// TIA Portal project "CLU" (V13) (continued)
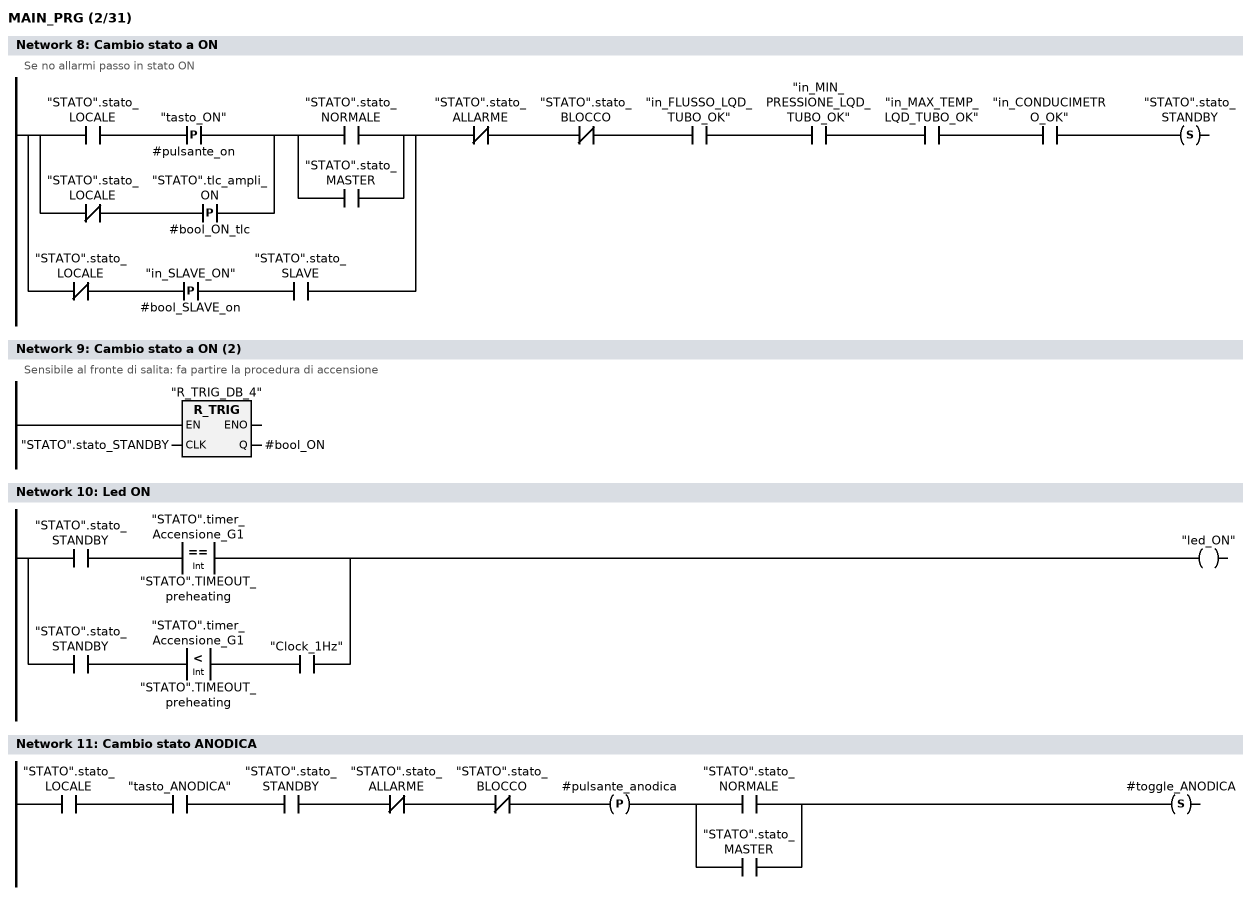
   RUNG wire#powerrail
      Contact( "STATO".stato_LOCALE )
      P_Contact(operand := "tasto_ON", bit := #pulsante_on)
      wire#w1
      Contact( "STATO".stato_NORMALE )
      wire#w2
      I_Contact( "STATO".stato_ALLARME )
      I_Contact( "STATO".stato_BLOCCO )
      Contact( "in_FLUSSO_LQD_TUBO_OK" )
      Contact( "in_MIN_PRESSIONE_LQD_TUBO_OK" )
      Contact( "in_MAX_TEMP_LQD_TUBO_OK" )
      Contact( "in_CONDUCIMETRO_OK" )
      S_Coil( "STATO".stato_STANDBY )
   END_RUNG
   RUNG wire#powerrail
      I_Contact( "STATO".stato_LOCALE )
      P_Contact(operand := "STATO".tlc_ampli_ON, bit := #bool_ON_tlc)
   END_RUNG wire#w1
   RUNG wire#w1
      Contact( "STATO".stato_MASTER )
   END_RUNG wire#w2
   RUNG wire#powerrail
      I_Contact( "STATO".stato_LOCALE )
      P_Contact(operand := "in_SLAVE_ON", bit := #bool_SLAVE_on)
      Contact( "STATO".stato_SLAVE )
   END_RUNG wire#w2
   // the same network as SCL:
   #_w1 := "STATO".stato_LOCALE AND "tasto_ON" AND NOT #pulsante_on;   // rising edge of "tasto_ON"
   #pulsante_on := "tasto_ON";
   #_w2 := NOT "STATO".stato_LOCALE AND "STATO".tlc_ampli_ON AND NOT #bool_ON_tlc;   // rising edge of "STATO".tlc_ampli_ON
   #bool_ON_tlc := "STATO".tlc_ampli_ON;
   #_w3 := NOT "STATO".stato_LOCALE AND "in_SLAVE_ON" AND NOT #bool_SLAVE_on;   // rising edge of "in_SLAVE_ON"
   #bool_SLAVE_on := "in_SLAVE_ON";
   IF (((#_w1 OR #_w2) AND ("STATO".stato_NORMALE OR "STATO".stato_MASTER)) OR (#_w3 AND "STATO".stato_SLAVE)) AND NOT "STATO".stato_ALLARME AND NOT "STATO".stato_BLOCCO AND "in_FLUSSO_LQD_TUBO_OK" AND "in_MIN_PRESSIONE_LQD_TUBO_OK" AND "in_MAX_TEMP_LQD_TUBO_OK" AND "in_CONDUCIMETRO_OK" THEN
       "STATO".stato_STANDBY := TRUE;
   END_IF;
END_REGION

REGION Network 9: Cambio stato a ON (2)
   // Sensibile al fronte di salita: fa partire la procedura di accensione
   "R_TRIG_DB_4"(CLK := "STATO".stato_STANDBY, Q => #bool_ON);   // R_TRIG
END_REGION

REGION Network 10: Led ON
   RUNG wire#powerrail
      Contact( "STATO".stato_STANDBY )
      { S7_Templates := "SrcType := Int" } EQ_Contact(in1 := "STATO".timer_Accensione_G1, in2 := "STATO".TIMEOUT_preheating)
      wire#w1
      Coil( "led_ON" )
   END_RUNG
   RUNG wire#powerrail
      Contact( "STATO".stato_STANDBY )
      { S7_Templates := "SrcType := Int" } LT_Contact(in1 := "STATO".timer_Accensione_G1, in2 := "STATO".TIMEOUT_preheating)
      Contact( "Clock_1Hz" )
   END_RUNG wire#w1
   // the same network as SCL:
   "led_ON" := ("STATO".stato_STANDBY AND ("STATO".timer_Accensione_G1 = "STATO".TIMEOUT_preheating)) OR ("STATO".stato_STANDBY AND ("STATO".timer_Accensione_G1 < "STATO".TIMEOUT_preheating) AND "Clock_1Hz");
END_REGION

REGION Network 11: Cambio stato ANODICA
   RUNG wire#powerrail
      Contact( "STATO".stato_LOCALE )
      Contact( "tasto_ANODICA" )
      Contact( "STATO".stato_STANDBY )
      I_Contact( "STATO".stato_ALLARME )
      I_Contact( "STATO".stato_BLOCCO )
      P_Trig( #pulsante_anodica )
      wire#w1
      Contact( "STATO".stato_NORMALE )
      wire#w2
      S_Coil( #toggle_ANODICA )
   END_RUNG
   RUNG wire#w1
      Contact( "STATO".stato_MASTER )
   END_RUNG wire#w2
   // the same network as SCL:
   #_w1 := "STATO".stato_LOCALE AND "tasto_ANODICA" AND "STATO".stato_STANDBY AND NOT "STATO".stato_ALLARME AND NOT "STATO".stato_BLOCCO;
   #_w2 := #_w1 AND NOT #pulsante_anodica;   // rising edge
   #pulsante_anodica := #_w1;
   IF #_w2 AND ("STATO".stato_NORMALE OR "STATO".stato_MASTER) THEN #toggle_ANODICA := TRUE; END_IF;
END_REGION

REGION Network 12: ANODICA ON
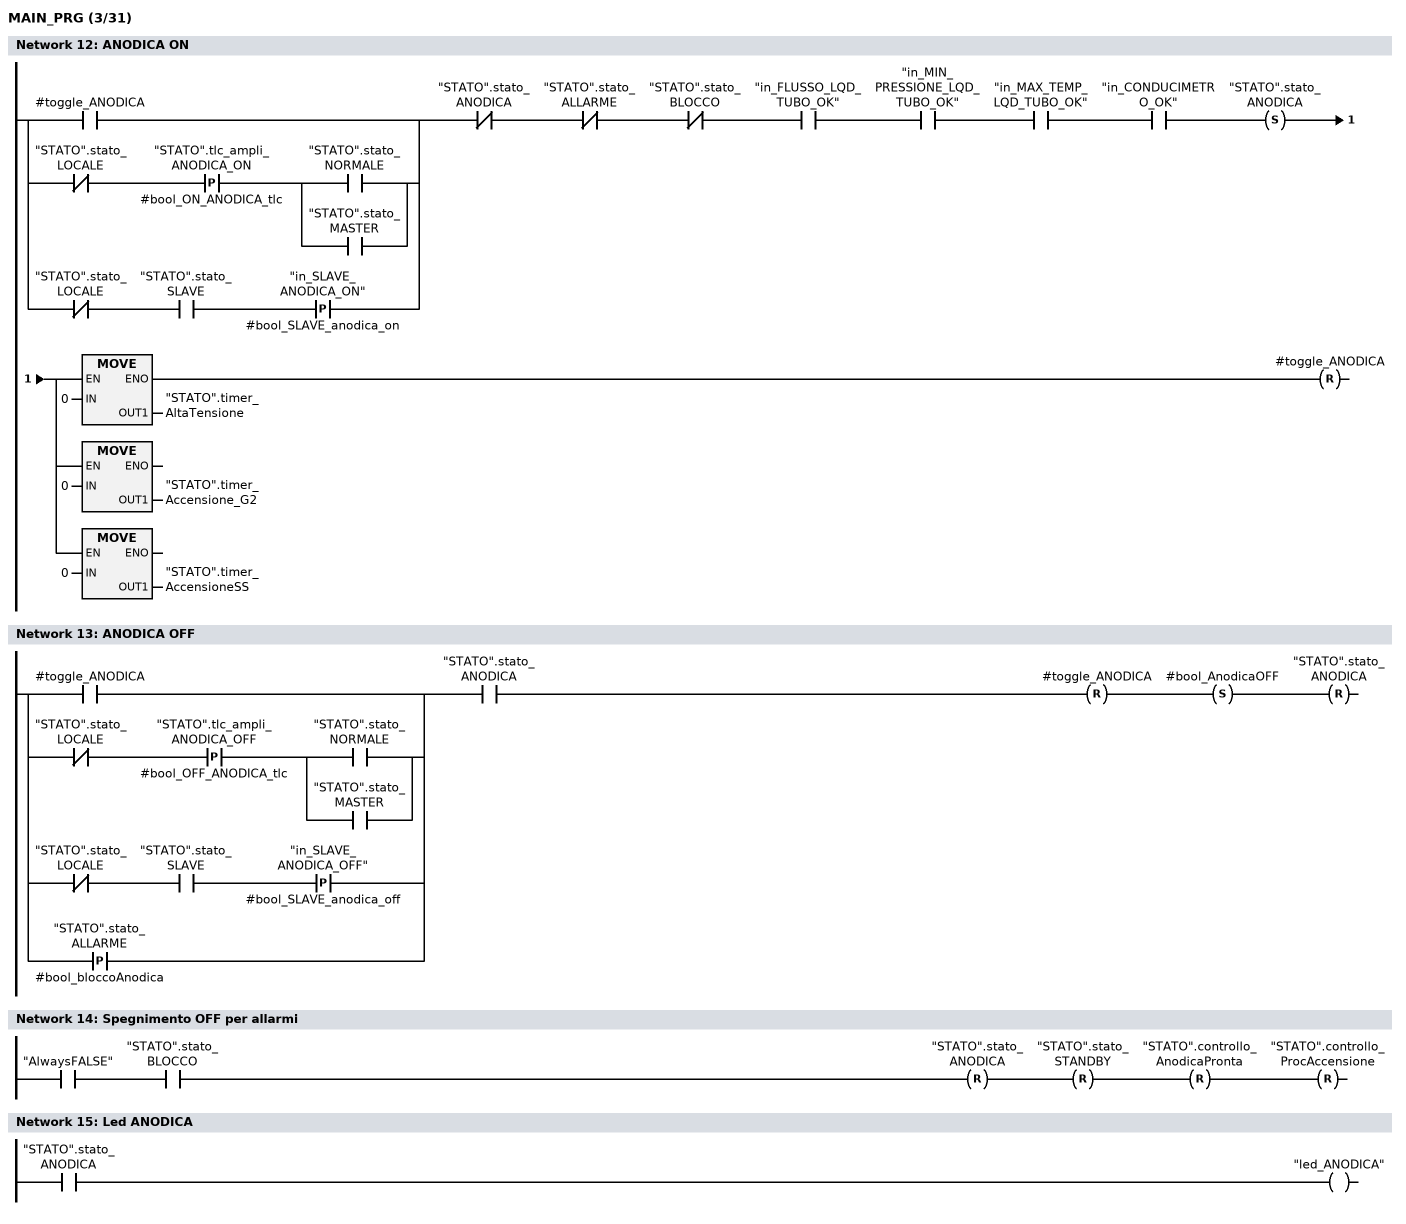
   RUNG wire#powerrail
      Contact( #toggle_ANODICA )
      wire#w1
      I_Contact( "STATO".stato_ANODICA )
      I_Contact( "STATO".stato_ALLARME )
      I_Contact( "STATO".stato_BLOCCO )
      Contact( "in_FLUSSO_LQD_TUBO_OK" )
      Contact( "in_MIN_PRESSIONE_LQD_TUBO_OK" )
      Contact( "in_MAX_TEMP_LQD_TUBO_OK" )
      Contact( "in_CONDUCIMETRO_OK" )
      S_Coil( "STATO".stato_ANODICA )
      wire#w3
      Move(in := 0, out1 => "STATO".timer_AltaTensione)
      R_Coil( #toggle_ANODICA )
   END_RUNG
   RUNG wire#powerrail
      I_Contact( "STATO".stato_LOCALE )
      P_Contact(operand := "STATO".tlc_ampli_ANODICA_ON, bit := #bool_ON_ANODICA_tlc)
      wire#w2
      Contact( "STATO".stato_NORMALE )
   END_RUNG wire#w1
   RUNG wire#w2
      Contact( "STATO".stato_MASTER )
   END_RUNG wire#w1
   RUNG wire#powerrail
      I_Contact( "STATO".stato_LOCALE )
      Contact( "STATO".stato_SLAVE )
      P_Contact(operand := "in_SLAVE_ANODICA_ON", bit := #bool_SLAVE_anodica_on)
   END_RUNG wire#w1
   RUNG wire#w3
      Move(in := 0, out1 => "STATO".timer_Accensione_G2)
   END_RUNG
   RUNG wire#w3
      Move(in := 0, out1 => "STATO".timer_AccensioneSS)
   END_RUNG
   // the same network as SCL:
   #_w1 := NOT "STATO".stato_LOCALE AND "STATO".tlc_ampli_ANODICA_ON AND NOT #bool_ON_ANODICA_tlc;   // rising edge of "STATO".tlc_ampli_ANODICA_ON
   #bool_ON_ANODICA_tlc := "STATO".tlc_ampli_ANODICA_ON;
   #_w2 := NOT "STATO".stato_LOCALE AND "STATO".stato_SLAVE AND "in_SLAVE_ANODICA_ON" AND NOT #bool_SLAVE_anodica_on;   // rising edge of "in_SLAVE_ANODICA_ON"
   #bool_SLAVE_anodica_on := "in_SLAVE_ANODICA_ON";
   #_w3 := (#toggle_ANODICA OR (#_w1 AND ("STATO".stato_NORMALE OR "STATO".stato_MASTER)) OR #_w2) AND NOT "STATO".stato_ANODICA AND NOT "STATO".stato_ALLARME AND NOT "STATO".stato_BLOCCO AND "in_FLUSSO_LQD_TUBO_OK" AND "in_MIN_PRESSIONE_LQD_TUBO_OK" AND "in_MAX_TEMP_LQD_TUBO_OK" AND "in_CONDUCIMETRO_OK";
   IF #_w3 THEN
       "STATO".stato_ANODICA := TRUE;
       "STATO".timer_AltaTensione := 0;
       #toggle_ANODICA := FALSE;
       "STATO".timer_Accensione_G2 := 0;
       "STATO".timer_AccensioneSS := 0;
   END_IF;
END_REGION

REGION Network 13: ANODICA OFF
   RUNG wire#powerrail
      Contact( #toggle_ANODICA )
      wire#w1
      Contact( "STATO".stato_ANODICA )
      R_Coil( #toggle_ANODICA )
      S_Coil( #bool_AnodicaOFF )
      R_Coil( "STATO".stato_ANODICA )
   END_RUNG
   RUNG wire#powerrail
      I_Contact( "STATO".stato_LOCALE )
      P_Contact(operand := "STATO".tlc_ampli_ANODICA_OFF, bit := #bool_OFF_ANODICA_tlc)
      wire#w2
      Contact( "STATO".stato_NORMALE )
   END_RUNG wire#w1
   RUNG wire#w2
      Contact( "STATO".stato_MASTER )
   END_RUNG wire#w1
   RUNG wire#powerrail
      I_Contact( "STATO".stato_LOCALE )
      Contact( "STATO".stato_SLAVE )
      P_Contact(operand := "in_SLAVE_ANODICA_OFF", bit := #bool_SLAVE_anodica_off)
   END_RUNG wire#w1
   RUNG wire#powerrail
      P_Contact(operand := "STATO".stato_ALLARME, bit := #bool_bloccoAnodica)
   END_RUNG wire#w1
   // the same network as SCL:
   #_w1 := NOT "STATO".stato_LOCALE AND "STATO".tlc_ampli_ANODICA_OFF AND NOT #bool_OFF_ANODICA_tlc;   // rising edge of "STATO".tlc_ampli_ANODICA_OFF
   #bool_OFF_ANODICA_tlc := "STATO".tlc_ampli_ANODICA_OFF;
   #_w2 := NOT "STATO".stato_LOCALE AND "STATO".stato_SLAVE AND "in_SLAVE_ANODICA_OFF" AND NOT #bool_SLAVE_anodica_off;   // rising edge of "in_SLAVE_ANODICA_OFF"
   #bool_SLAVE_anodica_off := "in_SLAVE_ANODICA_OFF";
   #_w3 := "STATO".stato_ALLARME AND NOT #bool_bloccoAnodica;   // rising edge of "STATO".stato_ALLARME
   #bool_bloccoAnodica := "STATO".stato_ALLARME;
   #_w4 := (#toggle_ANODICA OR (#_w1 AND ("STATO".stato_NORMALE OR "STATO".stato_MASTER)) OR #_w2 OR #_w3) AND "STATO".stato_ANODICA;
   IF #_w4 THEN
       #toggle_ANODICA := FALSE;
       #bool_AnodicaOFF := TRUE;
       "STATO".stato_ANODICA := FALSE;
   END_IF;
END_REGION

REGION Network 14: Spegnimento OFF per allarmi
   RUNG wire#powerrail
      Contact( "AlwaysFALSE" )
      Contact( "STATO".stato_BLOCCO )
      R_Coil( "STATO".stato_ANODICA )
      R_Coil( "STATO".stato_STANDBY )
      R_Coil( "STATO".controllo_AnodicaPronta )
      R_Coil( "STATO".controllo_ProcAccensione )
   END_RUNG
   // the same network as SCL:
   IF "AlwaysFALSE" AND "STATO".stato_BLOCCO THEN
       "STATO".stato_ANODICA := FALSE;
       "STATO".stato_STANDBY := FALSE;
       "STATO".controllo_AnodicaPronta := FALSE;
       "STATO".controllo_ProcAccensione := FALSE;
   END_IF;
END_REGION

REGION Network 15: Led ANODICA
   RUNG wire#powerrail
      Contact( "STATO".stato_ANODICA )
      Coil( "led_ANODICA" )
   END_RUNG
   // the same network as SCL:
   "led_ANODICA" := "STATO".stato_ANODICA;
END_REGION

REGION Network 16: Cambio a modo CW /Pulsed
   // Non applicabile se l'Anodica è attiva
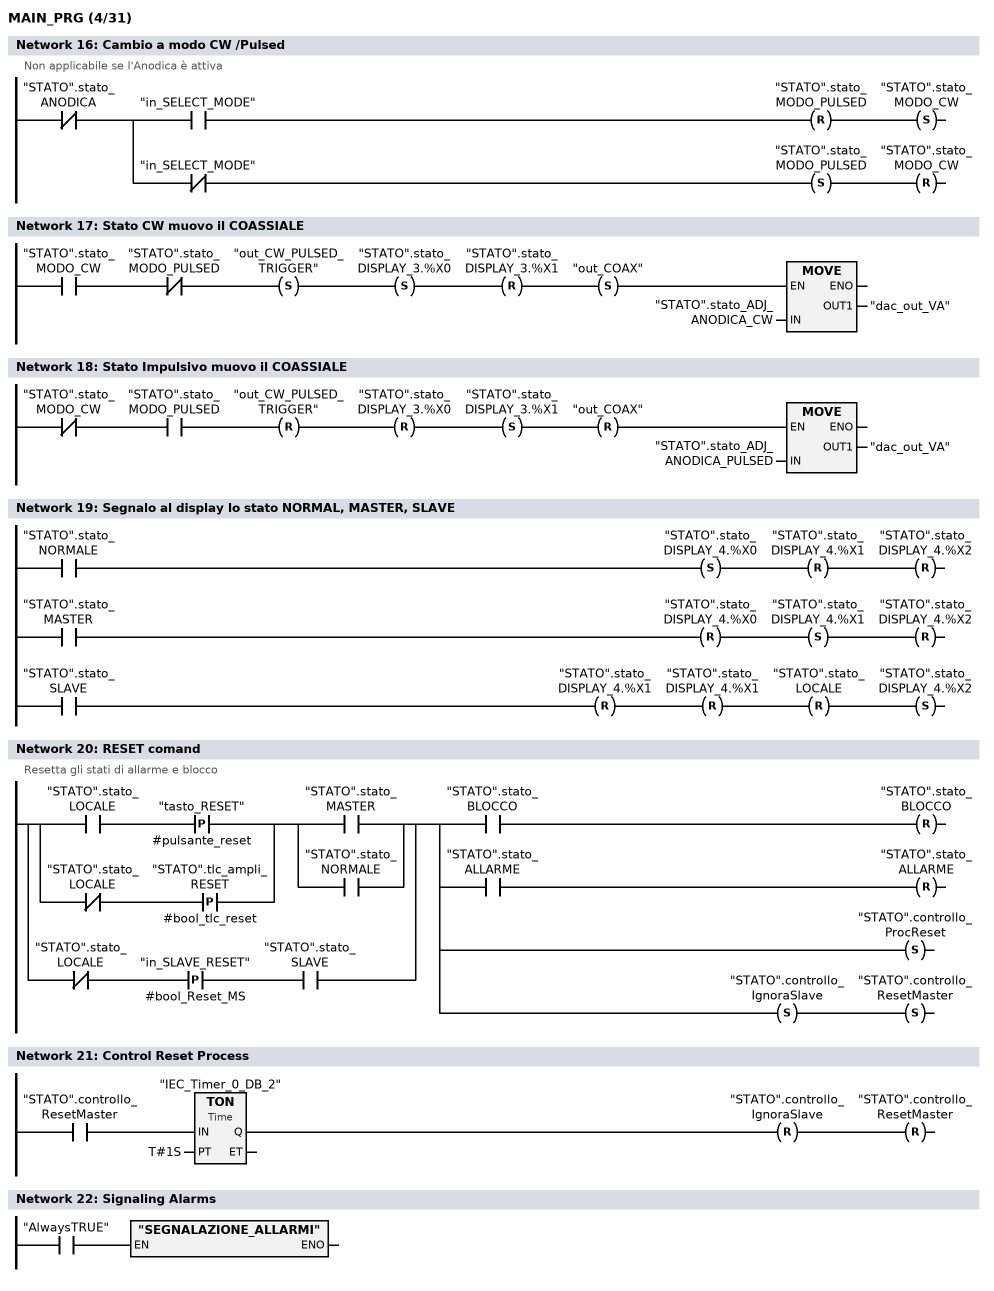
   RUNG wire#powerrail
      I_Contact( "STATO".stato_ANODICA )
      wire#w1
      Contact( "in_SELECT_MODE" )
      R_Coil( "STATO".stato_MODO_PULSED )
      S_Coil( "STATO".stato_MODO_CW )
   END_RUNG
   RUNG wire#w1
      I_Contact( "in_SELECT_MODE" )
      S_Coil( "STATO".stato_MODO_PULSED )
      R_Coil( "STATO".stato_MODO_CW )
   END_RUNG
   // the same network as SCL:
   #_w1 := NOT "STATO".stato_ANODICA;
   IF #_w1 AND "in_SELECT_MODE" THEN
       "STATO".stato_MODO_PULSED := FALSE;
       "STATO".stato_MODO_CW := TRUE;
   END_IF;
   IF #_w1 AND NOT "in_SELECT_MODE" THEN
       "STATO".stato_MODO_PULSED := TRUE;
       "STATO".stato_MODO_CW := FALSE;
   END_IF;
END_REGION

REGION Network 17: Stato CW muovo il COASSIALE
   RUNG wire#powerrail
      Contact( "STATO".stato_MODO_CW )
      I_Contact( "STATO".stato_MODO_PULSED )
      S_Coil( "out_CW_PULSED_TRIGGER" )
      S_Coil( "STATO".stato_DISPLAY_3.%X0 )
      R_Coil( "STATO".stato_DISPLAY_3.%X1 )
      S_Coil( "out_COAX" )
      Move(in := "STATO".stato_ADJ_ANODICA_CW, out1 => "dac_out_VA")
   END_RUNG
   // the same network as SCL:
   IF "STATO".stato_MODO_CW AND NOT "STATO".stato_MODO_PULSED THEN
       "out_CW_PULSED_TRIGGER" := TRUE;
       "STATO".stato_DISPLAY_3.%X0 := TRUE;
       "STATO".stato_DISPLAY_3.%X1 := FALSE;
       "out_COAX" := TRUE;
       "dac_out_VA" := "STATO".stato_ADJ_ANODICA_CW;
   END_IF;
END_REGION

REGION Network 18: Stato Impulsivo muovo il COASSIALE
   RUNG wire#powerrail
      I_Contact( "STATO".stato_MODO_CW )
      Contact( "STATO".stato_MODO_PULSED )
      R_Coil( "out_CW_PULSED_TRIGGER" )
      R_Coil( "STATO".stato_DISPLAY_3.%X0 )
      S_Coil( "STATO".stato_DISPLAY_3.%X1 )
      R_Coil( "out_COAX" )
      Move(in := "STATO".stato_ADJ_ANODICA_PULSED, out1 => "dac_out_VA")
   END_RUNG
   // the same network as SCL:
   IF NOT "STATO".stato_MODO_CW AND "STATO".stato_MODO_PULSED THEN
       "out_CW_PULSED_TRIGGER" := FALSE;
       "STATO".stato_DISPLAY_3.%X0 := FALSE;
       "STATO".stato_DISPLAY_3.%X1 := TRUE;
       "out_COAX" := FALSE;
       "dac_out_VA" := "STATO".stato_ADJ_ANODICA_PULSED;
   END_IF;
END_REGION

REGION Network 19: Segnalo al display lo stato NORMAL, MASTER, SLAVE
   RUNG wire#powerrail
      Contact( "STATO".stato_NORMALE )
      S_Coil( "STATO".stato_DISPLAY_4.%X0 )
      R_Coil( "STATO".stato_DISPLAY_4.%X1 )
      R_Coil( "STATO".stato_DISPLAY_4.%X2 )
   END_RUNG
   RUNG wire#powerrail
      Contact( "STATO".stato_MASTER )
      R_Coil( "STATO".stato_DISPLAY_4.%X0 )
      S_Coil( "STATO".stato_DISPLAY_4.%X1 )
      R_Coil( "STATO".stato_DISPLAY_4.%X2 )
   END_RUNG
   RUNG wire#powerrail
      Contact( "STATO".stato_SLAVE )
      R_Coil( "STATO".stato_DISPLAY_4.%X1 )
      R_Coil( "STATO".stato_DISPLAY_4.%X1 )
      R_Coil( "STATO".stato_LOCALE )
      S_Coil( "STATO".stato_DISPLAY_4.%X2 )
   END_RUNG
   // the same network as SCL:
   IF "STATO".stato_NORMALE THEN
       "STATO".stato_DISPLAY_4.%X0 := TRUE;
       "STATO".stato_DISPLAY_4.%X1 := FALSE;
       "STATO".stato_DISPLAY_4.%X2 := FALSE;
   END_IF;
   IF "STATO".stato_MASTER THEN
       "STATO".stato_DISPLAY_4.%X0 := FALSE;
       "STATO".stato_DISPLAY_4.%X1 := TRUE;
       "STATO".stato_DISPLAY_4.%X2 := FALSE;
   END_IF;
   IF "STATO".stato_SLAVE THEN
       "STATO".stato_DISPLAY_4.%X1 := FALSE;
       "STATO".stato_DISPLAY_4.%X1 := FALSE;
       "STATO".stato_LOCALE := FALSE;
       "STATO".stato_DISPLAY_4.%X2 := TRUE;
   END_IF;
END_REGION

REGION Network 20: RESET comand
   // Resetta gli stati di allarme e blocco
   RUNG wire#powerrail
      Contact( "STATO".stato_LOCALE )
      P_Contact(operand := "tasto_RESET", bit := #pulsante_reset)
      wire#w1
      Contact( "STATO".stato_MASTER )
      wire#w2
      Contact( "STATO".stato_BLOCCO )
      R_Coil( "STATO".stato_BLOCCO )
   END_RUNG
   RUNG wire#powerrail
      I_Contact( "STATO".stato_LOCALE )
      P_Contact(operand := "STATO".tlc_ampli_RESET, bit := #bool_tlc_reset)
   END_RUNG wire#w1
   RUNG wire#w1
      Contact( "STATO".stato_NORMALE )
   END_RUNG wire#w2
   RUNG wire#powerrail
      I_Contact( "STATO".stato_LOCALE )
      P_Contact(operand := "in_SLAVE_RESET", bit := #bool_Reset_MS)
      Contact( "STATO".stato_SLAVE )
   END_RUNG wire#w2
   RUNG wire#w2
      Contact( "STATO".stato_ALLARME )
      R_Coil( "STATO".stato_ALLARME )
   END_RUNG
   RUNG wire#w2
      S_Coil( "STATO".controllo_ProcReset )
   END_RUNG
   RUNG wire#w2
      S_Coil( "STATO".controllo_IgnoraSlave )
      S_Coil( "STATO".controllo_ResetMaster )
   END_RUNG
   // the same network as SCL:
   #_w1 := "STATO".stato_LOCALE AND "tasto_RESET" AND NOT #pulsante_reset;   // rising edge of "tasto_RESET"
   #pulsante_reset := "tasto_RESET";
   #_w2 := NOT "STATO".stato_LOCALE AND "STATO".tlc_ampli_RESET AND NOT #bool_tlc_reset;   // rising edge of "STATO".tlc_ampli_RESET
   #bool_tlc_reset := "STATO".tlc_ampli_RESET;
   #_w3 := NOT "STATO".stato_LOCALE AND "in_SLAVE_RESET" AND NOT #bool_Reset_MS;   // rising edge of "in_SLAVE_RESET"
   #bool_Reset_MS := "in_SLAVE_RESET";
   #_w4 := ((#_w1 OR #_w2) AND ("STATO".stato_MASTER OR "STATO".stato_NORMALE)) OR (#_w3 AND "STATO".stato_SLAVE);
   IF #_w4 AND "STATO".stato_BLOCCO THEN "STATO".stato_BLOCCO := FALSE; END_IF;
   IF #_w4 AND "STATO".stato_ALLARME THEN "STATO".stato_ALLARME := FALSE; END_IF;
   IF #_w4 THEN
       "STATO".controllo_ProcReset := TRUE;
       "STATO".controllo_IgnoraSlave := TRUE;
       "STATO".controllo_ResetMaster := TRUE;
   END_IF;
END_REGION

REGION Network 21: Control Reset Process
   "IEC_Timer_0_DB_2".TON(IN := "STATO".controllo_ResetMaster, PT := T#1S);
   IF "IEC_Timer_0_DB_2".Q THEN
       "STATO".controllo_IgnoraSlave := FALSE;
       "STATO".controllo_ResetMaster := FALSE;
   END_IF;
END_REGION

REGION Network 22: Signaling Alarms
   RUNG wire#powerrail
      Contact( "AlwaysTRUE" )
      "SEGNALAZIONE_ALLARMI"()
   END_RUNG
   // the same network as SCL:
   IF "AlwaysTRUE" THEN "SEGNALAZIONE_ALLARMI"(); END_IF;
END_REGION

REGION Network 23: Erasing Alarms
   // In seguito ad un reset.
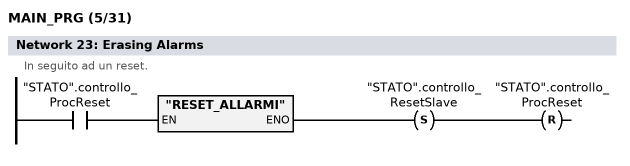
   RUNG wire#powerrail
      Contact( "STATO".controllo_ProcReset )
      "RESET_ALLARMI"()
      S_Coil( "STATO".controllo_ResetSlave )
      R_Coil( "STATO".controllo_ProcReset )
   END_RUNG
   // the same network as SCL:
   "RESET_ALLARMI"(EN := "STATO".controllo_ProcReset, ENO => #_w1);
   IF #_w1 THEN
       "STATO".controllo_ResetSlave := TRUE;
       "STATO".controllo_ProcReset := FALSE;
   END_IF;
END_REGION

REGION Network 24: ALARM STATE
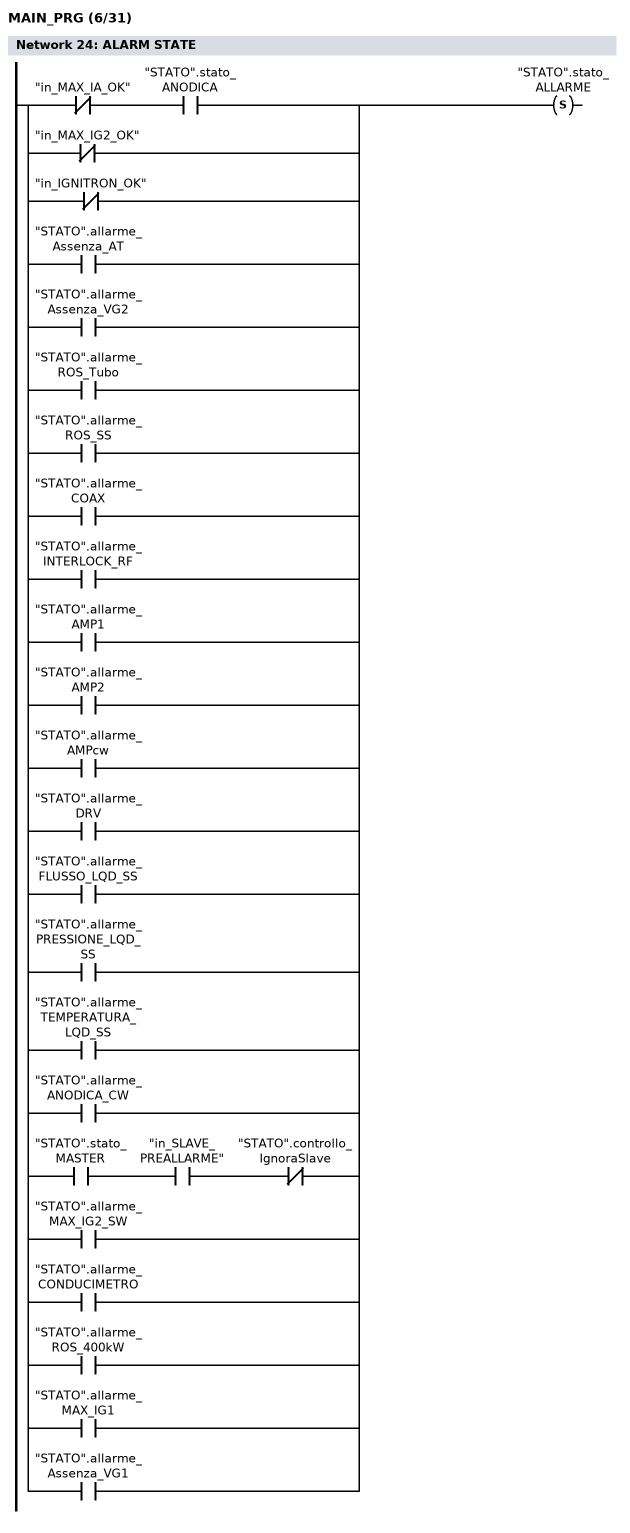
   RUNG wire#powerrail
      I_Contact( "in_MAX_IA_OK" )
      Contact( "STATO".stato_ANODICA )
      wire#w1
      S_Coil( "STATO".stato_ALLARME )
   END_RUNG
   RUNG wire#powerrail
      I_Contact( "in_MAX_IG2_OK" )
   END_RUNG wire#w1
   RUNG wire#powerrail
      I_Contact( "in_IGNITRON_OK" )
   END_RUNG wire#w1
   RUNG wire#powerrail
      Contact( "STATO".allarme_Assenza_AT )
   END_RUNG wire#w1
   RUNG wire#powerrail
      Contact( "STATO".allarme_Assenza_VG2 )
   END_RUNG wire#w1
   RUNG wire#powerrail
      Contact( "STATO".allarme_ROS_Tubo )
   END_RUNG wire#w1
   RUNG wire#powerrail
      Contact( "STATO".allarme_ROS_SS )
   END_RUNG wire#w1
   RUNG wire#powerrail
      Contact( "STATO".allarme_COAX )
   END_RUNG wire#w1
   RUNG wire#powerrail
      Contact( "STATO".allarme_INTERLOCK_RF )
   END_RUNG wire#w1
   RUNG wire#powerrail
      Contact( "STATO".allarme_AMP1 )
   END_RUNG wire#w1
   RUNG wire#powerrail
      Contact( "STATO".allarme_AMP2 )
   END_RUNG wire#w1
   RUNG wire#powerrail
      Contact( "STATO".allarme_AMPcw )
   END_RUNG wire#w1
   RUNG wire#powerrail
      Contact( "STATO".allarme_DRV )
   END_RUNG wire#w1
   RUNG wire#powerrail
      Contact( "STATO".allarme_FLUSSO_LQD_SS )
   END_RUNG wire#w1
   RUNG wire#powerrail
      Contact( "STATO".allarme_PRESSIONE_LQD_SS )
   END_RUNG wire#w1
   RUNG wire#powerrail
      Contact( "STATO".allarme_TEMPERATURA_LQD_SS )
   END_RUNG wire#w1
   RUNG wire#powerrail
      Contact( "STATO".allarme_ANODICA_CW )
   END_RUNG wire#w1
   RUNG wire#powerrail
      Contact( "STATO".stato_MASTER )
      Contact( "in_SLAVE_PREALLARME" )
      I_Contact( "STATO".controllo_IgnoraSlave )
   END_RUNG wire#w1
   RUNG wire#powerrail
      Contact( "STATO".allarme_MAX_IG2_SW )
   END_RUNG wire#w1
   RUNG wire#powerrail
      Contact( "STATO".allarme_CONDUCIMETRO )
   END_RUNG wire#w1
   RUNG wire#powerrail
      Contact( "STATO".allarme_ROS_400kW )
   END_RUNG wire#w1
   RUNG wire#powerrail
      Contact( "STATO".allarme_MAX_IG1 )
   END_RUNG wire#w1
   RUNG wire#powerrail
      Contact( "STATO".allarme_Assenza_VG1 )
   END_RUNG wire#w1
   // the same network as SCL:
   IF (NOT "in_MAX_IA_OK" AND "STATO".stato_ANODICA) OR NOT "in_MAX_IG2_OK" OR NOT "in_IGNITRON_OK" OR "STATO".allarme_Assenza_AT OR "STATO".allarme_Assenza_VG2 OR "STATO".allarme_ROS_Tubo OR "STATO".allarme_ROS_SS OR "STATO".allarme_COAX OR "STATO".allarme_INTERLOCK_RF OR "STATO".allarme_AMP1 OR "STATO".allarme_AMP2 OR "STATO".allarme_AMPcw OR "STATO".allarme_DRV OR "STATO".allarme_FLUSSO_LQD_SS OR "STATO".allarme_PRESSIONE_LQD_SS OR "STATO".allarme_TEMPERATURA_LQD_SS OR "STATO".allarme_ANODICA_CW OR ("STATO".stato_MASTER AND "in_SLAVE_PREALLARME" AND NOT "STATO".controllo_IgnoraSlave) OR "STATO".allarme_MAX_IG2_SW OR "STATO".allarme_CONDUCIMETRO OR "STATO".allarme_ROS_400kW OR "STATO".allarme_MAX_IG1 OR "STATO".allarme_Assenza_VG1 THEN
       "STATO".stato_ALLARME := TRUE;
   END_IF;
END_REGION

REGION Network 25: FAULT STATE
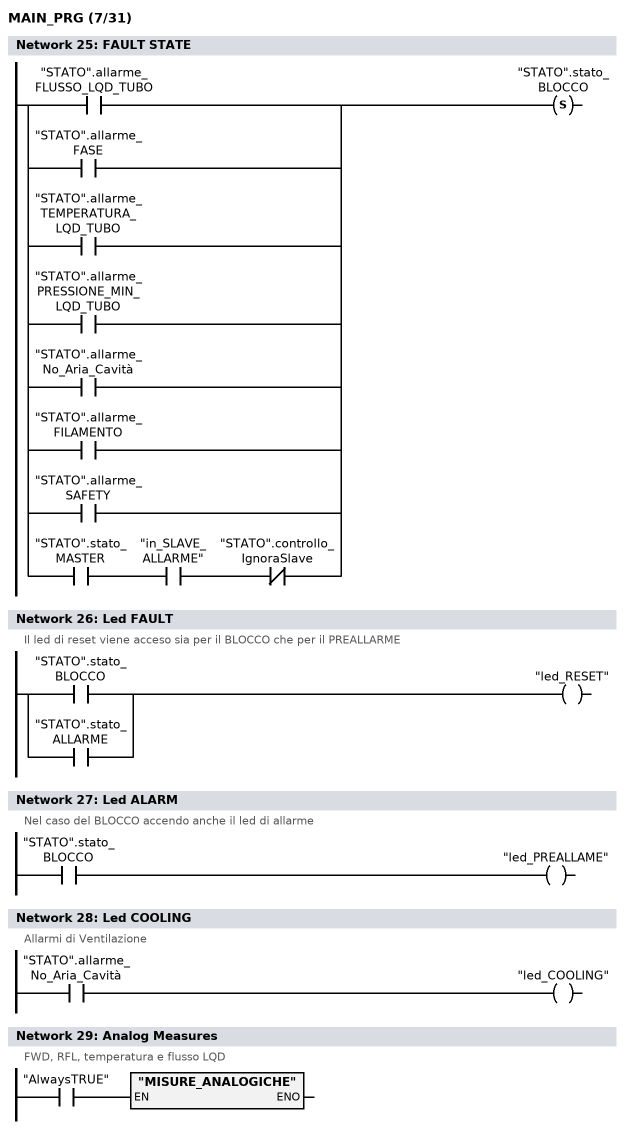
   RUNG wire#powerrail
      Contact( "STATO".allarme_FLUSSO_LQD_TUBO )
      wire#w1
      S_Coil( "STATO".stato_BLOCCO )
   END_RUNG
   RUNG wire#powerrail
      Contact( "STATO".allarme_FASE )
   END_RUNG wire#w1
   RUNG wire#powerrail
      Contact( "STATO".allarme_TEMPERATURA_LQD_TUBO )
   END_RUNG wire#w1
   RUNG wire#powerrail
      Contact( "STATO".allarme_PRESSIONE_MIN_LQD_TUBO )
   END_RUNG wire#w1
   RUNG wire#powerrail
      Contact( "STATO".allarme_No_Aria_Cavità )
   END_RUNG wire#w1
   RUNG wire#powerrail
      Contact( "STATO".allarme_FILAMENTO )
   END_RUNG wire#w1
   RUNG wire#powerrail
      Contact( "STATO".allarme_SAFETY )
   END_RUNG wire#w1
   RUNG wire#powerrail
      Contact( "STATO".stato_MASTER )
      Contact( "in_SLAVE_ALLARME" )
      I_Contact( "STATO".controllo_IgnoraSlave )
   END_RUNG wire#w1
   // the same network as SCL:
   IF "STATO".allarme_FLUSSO_LQD_TUBO OR "STATO".allarme_FASE OR "STATO".allarme_TEMPERATURA_LQD_TUBO OR "STATO".allarme_PRESSIONE_MIN_LQD_TUBO OR "STATO".allarme_No_Aria_Cavità OR "STATO".allarme_FILAMENTO OR "STATO".allarme_SAFETY OR ("STATO".stato_MASTER AND "in_SLAVE_ALLARME" AND NOT "STATO".controllo_IgnoraSlave) THEN
       "STATO".stato_BLOCCO := TRUE;
   END_IF;
END_REGION

REGION Network 26: Led FAULT
   // Il led di reset viene acceso sia per il BLOCCO che per il PREALLARME
   RUNG wire#powerrail
      Contact( "STATO".stato_BLOCCO )
      wire#w1
      Coil( "led_RESET" )
   END_RUNG
   RUNG wire#powerrail
      Contact( "STATO".stato_ALLARME )
   END_RUNG wire#w1
   // the same network as SCL:
   "led_RESET" := "STATO".stato_BLOCCO OR "STATO".stato_ALLARME;
END_REGION

REGION Network 27: Led ALARM
   // Nel caso del BLOCCO accendo anche il led di allarme
   RUNG wire#powerrail
      Contact( "STATO".stato_BLOCCO )
      Coil( "led_PREALLAME" )
   END_RUNG
   // the same network as SCL:
   "led_PREALLAME" := "STATO".stato_BLOCCO;
END_REGION

REGION Network 28: Led COOLING
   // Allarmi di Ventilazione
   RUNG wire#powerrail
      Contact( "STATO".allarme_No_Aria_Cavità )
      Coil( "led_COOLING" )
   END_RUNG
   // the same network as SCL:
   "led_COOLING" := "STATO".allarme_No_Aria_Cavità;
END_REGION

REGION Network 29: Analog Measures
   // FWD, RFL, temperatura e flusso LQD
   RUNG wire#powerrail
      Contact( "AlwaysTRUE" )
      "MISURE_ANALOGICHE"()
   END_RUNG
   // the same network as SCL:
   IF "AlwaysTRUE" THEN "MISURE_ANALOGICHE"(); END_IF;
END_REGION

REGION Network 30: PASSAGGIO IN STATO ON/STANDBY (1): start blowers
   // Inizio processo catena di accensione. Se non ci sono nallarmi attivo i ventilatori e inizializzo il timer accensione della griglia G1.